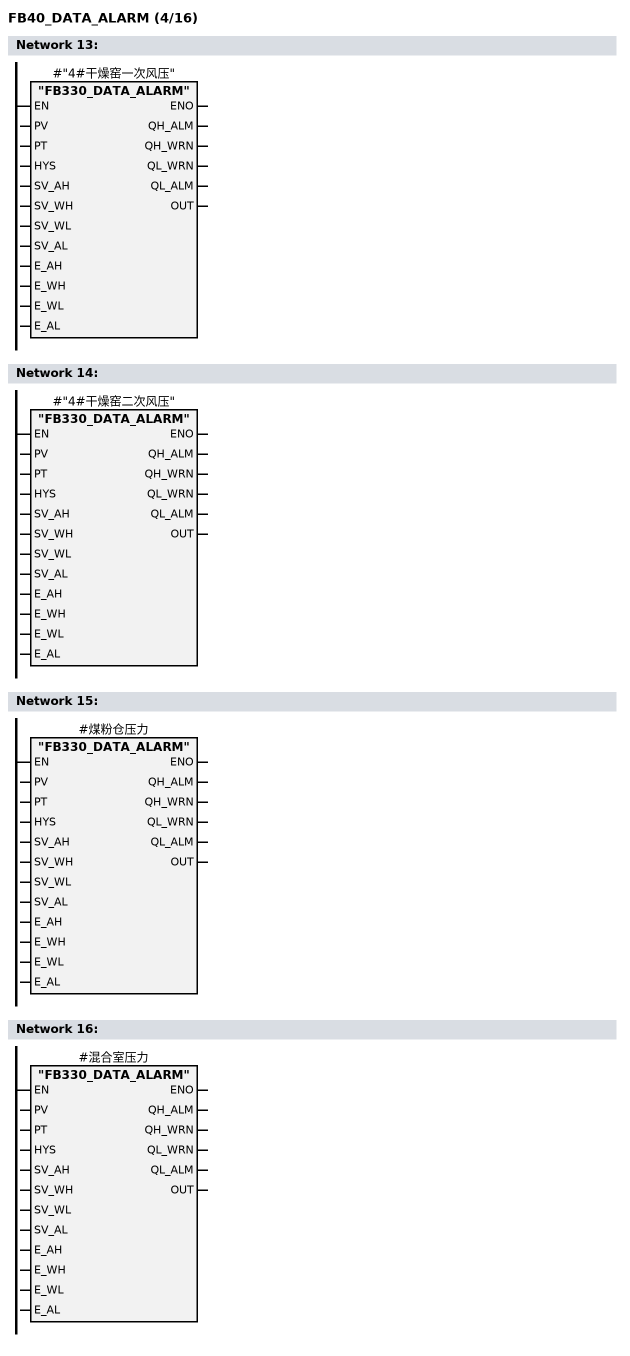
   RUNG wire#powerrail
      #"4#干燥窑一次风压"(PV :=, PT :=, HYS :=, SV_AH :=, SV_WH :=, SV_WL :=, SV_AL :=, E_AH :=, E_WH :=, E_WL :=, E_AL :=, QH_ALM =>, QH_WRN =>, QL_WRN =>, QL_ALM =>, OUT =>)
   END_RUNG
   // the same network as SCL:
   #"4#干燥窑一次风压"();   // "FB330_DATA_ALARM"
END_REGION

REGION Network 14
   RUNG wire#powerrail
      #"4#干燥窑二次风压"(PV :=, PT :=, HYS :=, SV_AH :=, SV_WH :=, SV_WL :=, SV_AL :=, E_AH :=, E_WH :=, E_WL :=, E_AL :=, QH_ALM =>, QH_WRN =>, QL_WRN =>, QL_ALM =>, OUT =>)
   END_RUNG
   // the same network as SCL:
   #"4#干燥窑二次风压"();   // "FB330_DATA_ALARM"
END_REGION

REGION Network 15
   RUNG wire#powerrail
      #煤粉仓压力(PV :=, PT :=, HYS :=, SV_AH :=, SV_WH :=, SV_WL :=, SV_AL :=, E_AH :=, E_WH :=, E_WL :=, E_AL :=, QH_ALM =>, QH_WRN =>, QL_WRN =>, QL_ALM =>, OUT =>)
   END_RUNG
   // the same network as SCL:
   #煤粉仓压力();   // "FB330_DATA_ALARM"
END_REGION

REGION Network 16
   RUNG wire#powerrail
      #混合室压力(PV :=, PT :=, HYS :=, SV_AH :=, SV_WH :=, SV_WL :=, SV_AL :=, E_AH :=, E_WH :=, E_WL :=, E_AL :=, QH_ALM =>, QH_WRN =>, QL_WRN =>, QL_ALM =>, OUT =>)
   END_RUNG
   // the same network as SCL:
   #混合室压力();   // "FB330_DATA_ALARM"
END_REGION

REGION Network 17
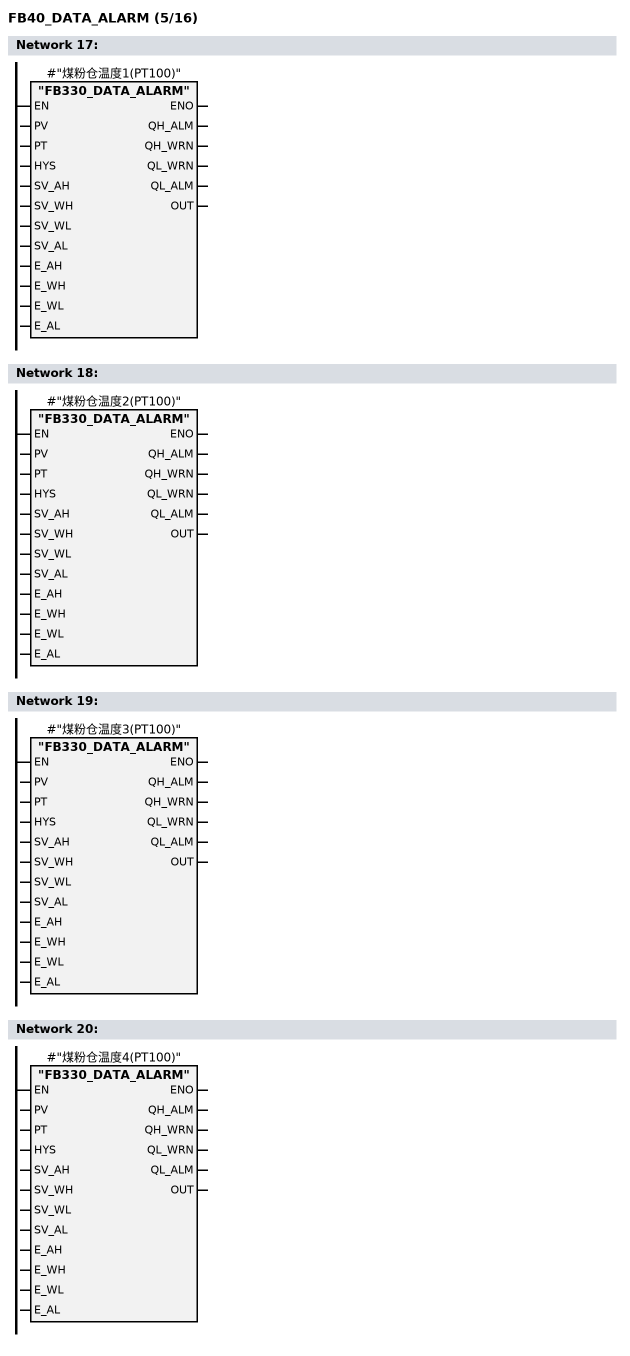
   RUNG wire#powerrail
      #"煤粉仓温度1(PT100)"(PV :=, PT :=, HYS :=, SV_AH :=, SV_WH :=, SV_WL :=, SV_AL :=, E_AH :=, E_WH :=, E_WL :=, E_AL :=, QH_ALM =>, QH_WRN =>, QL_WRN =>, QL_ALM =>, OUT =>)
   END_RUNG
   // the same network as SCL:
   #"煤粉仓温度1(PT100)"();   // "FB330_DATA_ALARM"
END_REGION

REGION Network 18
   RUNG wire#powerrail
      #"煤粉仓温度2(PT100)"(PV :=, PT :=, HYS :=, SV_AH :=, SV_WH :=, SV_WL :=, SV_AL :=, E_AH :=, E_WH :=, E_WL :=, E_AL :=, QH_ALM =>, QH_WRN =>, QL_WRN =>, QL_ALM =>, OUT =>)
   END_RUNG
   // the same network as SCL:
   #"煤粉仓温度2(PT100)"();   // "FB330_DATA_ALARM"
END_REGION

REGION Network 19
   RUNG wire#powerrail
      #"煤粉仓温度3(PT100)"(PV :=, PT :=, HYS :=, SV_AH :=, SV_WH :=, SV_WL :=, SV_AL :=, E_AH :=, E_WH :=, E_WL :=, E_AL :=, QH_ALM =>, QH_WRN =>, QL_WRN =>, QL_ALM =>, OUT =>)
   END_RUNG
   // the same network as SCL:
   #"煤粉仓温度3(PT100)"();   // "FB330_DATA_ALARM"
END_REGION

REGION Network 20
   RUNG wire#powerrail
      #"煤粉仓温度4(PT100)"(PV :=, PT :=, HYS :=, SV_AH :=, SV_WH :=, SV_WL :=, SV_AL :=, E_AH :=, E_WH :=, E_WL :=, E_AL :=, QH_ALM =>, QH_WRN =>, QL_WRN =>, QL_ALM =>, OUT =>)
   END_RUNG
   // the same network as SCL:
   #"煤粉仓温度4(PT100)"();   // "FB330_DATA_ALARM"
END_REGION

REGION Network 21
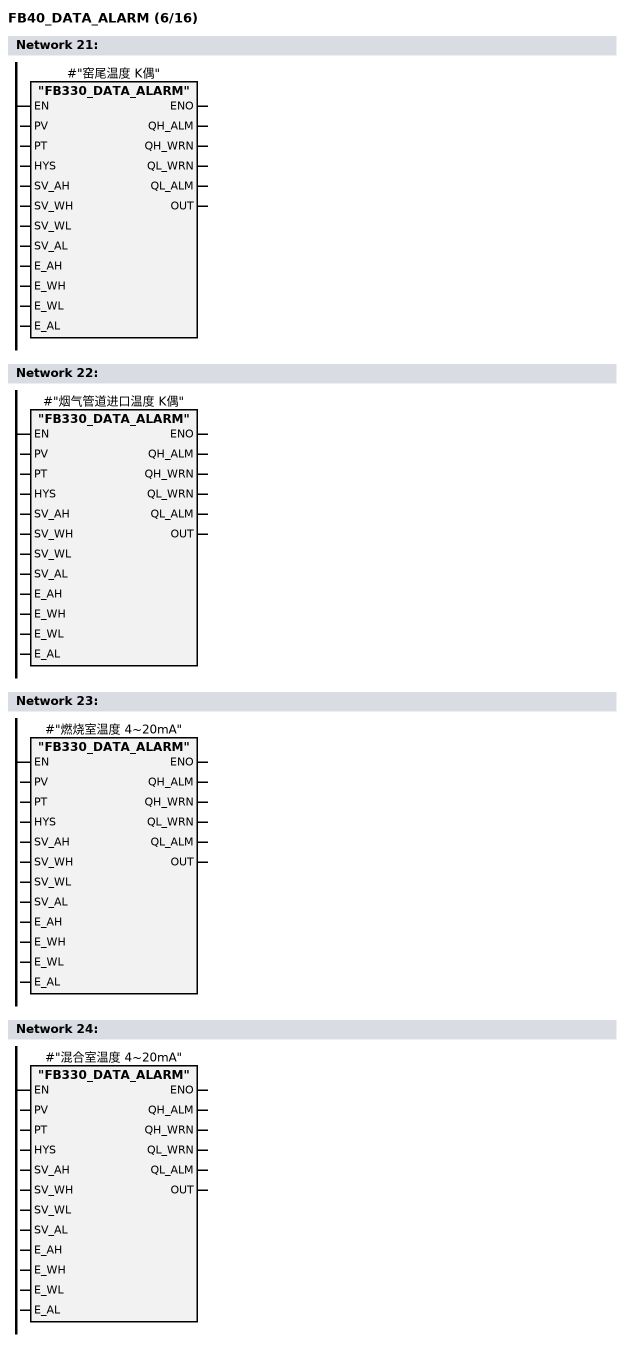
   RUNG wire#powerrail
      #"窑尾温度 K偶"(PV :=, PT :=, HYS :=, SV_AH :=, SV_WH :=, SV_WL :=, SV_AL :=, E_AH :=, E_WH :=, E_WL :=, E_AL :=, QH_ALM =>, QH_WRN =>, QL_WRN =>, QL_ALM =>, OUT =>)
   END_RUNG
   // the same network as SCL:
   #"窑尾温度 K偶"();   // "FB330_DATA_ALARM"
END_REGION

REGION Network 22
   RUNG wire#powerrail
      #"烟气管道进口温度 K偶"(PV :=, PT :=, HYS :=, SV_AH :=, SV_WH :=, SV_WL :=, SV_AL :=, E_AH :=, E_WH :=, E_WL :=, E_AL :=, QH_ALM =>, QH_WRN =>, QL_WRN =>, QL_ALM =>, OUT =>)
   END_RUNG
   // the same network as SCL:
   #"烟气管道进口温度 K偶"();   // "FB330_DATA_ALARM"
END_REGION

REGION Network 23
   RUNG wire#powerrail
      #"燃烧室温度 4~20mA"(PV :=, PT :=, HYS :=, SV_AH :=, SV_WH :=, SV_WL :=, SV_AL :=, E_AH :=, E_WH :=, E_WL :=, E_AL :=, QH_ALM =>, QH_WRN =>, QL_WRN =>, QL_ALM =>, OUT =>)
   END_RUNG
   // the same network as SCL:
   #"燃烧室温度 4~20mA"();   // "FB330_DATA_ALARM"
END_REGION

REGION Network 24
   RUNG wire#powerrail
      #"混合室温度 4~20mA"(PV :=, PT :=, HYS :=, SV_AH :=, SV_WH :=, SV_WL :=, SV_AL :=, E_AH :=, E_WH :=, E_WL :=, E_AL :=, QH_ALM =>, QH_WRN =>, QL_WRN =>, QL_ALM =>, OUT =>)
   END_RUNG
   // the same network as SCL:
   #"混合室温度 4~20mA"();   // "FB330_DATA_ALARM"
END_REGION

REGION Network 25
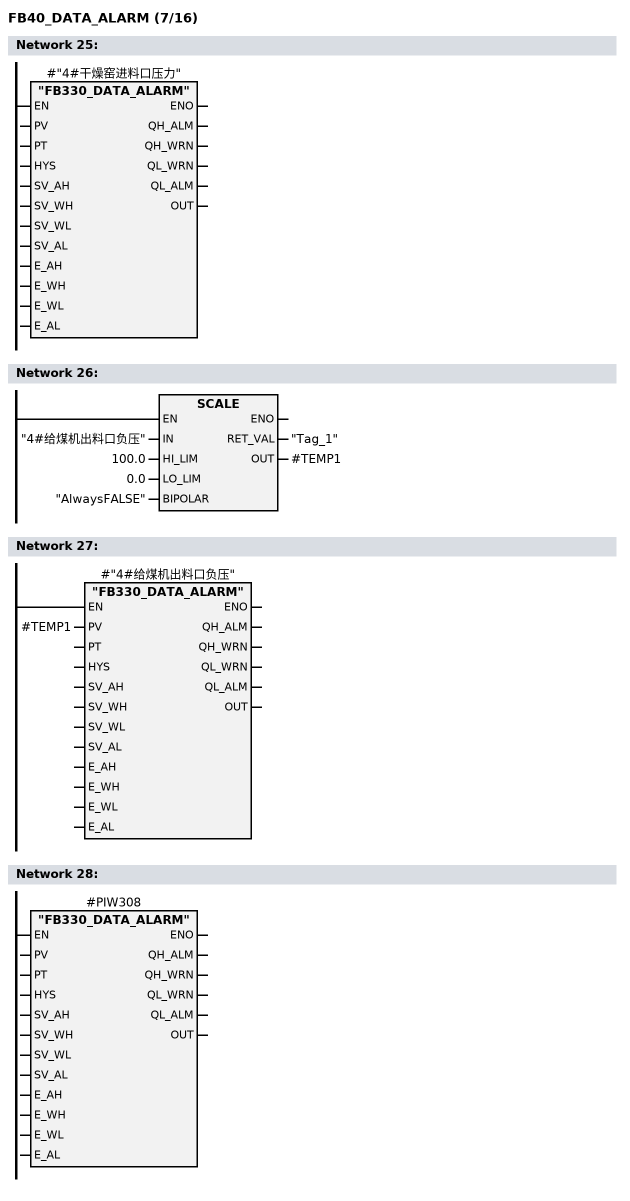
   RUNG wire#powerrail
      #"4#干燥窑进料口压力"(PV :=, PT :=, HYS :=, SV_AH :=, SV_WH :=, SV_WL :=, SV_AL :=, E_AH :=, E_WH :=, E_WL :=, E_AL :=, QH_ALM =>, QH_WRN =>, QL_WRN =>, QL_ALM =>, OUT =>)
   END_RUNG
   // the same network as SCL:
   #"4#干燥窑进料口压力"();   // "FB330_DATA_ALARM"
END_REGION

REGION Network 26
   "Tag_1" := SCALE(IN := "4#给煤机出料口负压", HI_LIM := 100.0, LO_LIM := 0.0, BIPOLAR := "AlwaysFALSE", OUT => #TEMP1);
END_REGION

REGION Network 27
   RUNG wire#powerrail
      #"4#给煤机出料口负压"(PV := #TEMP1, PT :=, HYS :=, SV_AH :=, SV_WH :=, SV_WL :=, SV_AL :=, E_AH :=, E_WH :=, E_WL :=, E_AL :=, QH_ALM =>, QH_WRN =>, QL_WRN =>, QL_ALM =>, OUT =>)
   END_RUNG
   // the same network as SCL:
   #"4#给煤机出料口负压"(PV := #TEMP1);   // "FB330_DATA_ALARM"
END_REGION

REGION Network 28
   RUNG wire#powerrail
      #PIW308(PV :=, PT :=, HYS :=, SV_AH :=, SV_WH :=, SV_WL :=, SV_AL :=, E_AH :=, E_WH :=, E_WL :=, E_AL :=, QH_ALM =>, QH_WRN =>, QL_WRN =>, QL_ALM =>, OUT =>)
   END_RUNG
   // the same network as SCL:
   #PIW308();   // "FB330_DATA_ALARM"
END_REGION

REGION Network 29
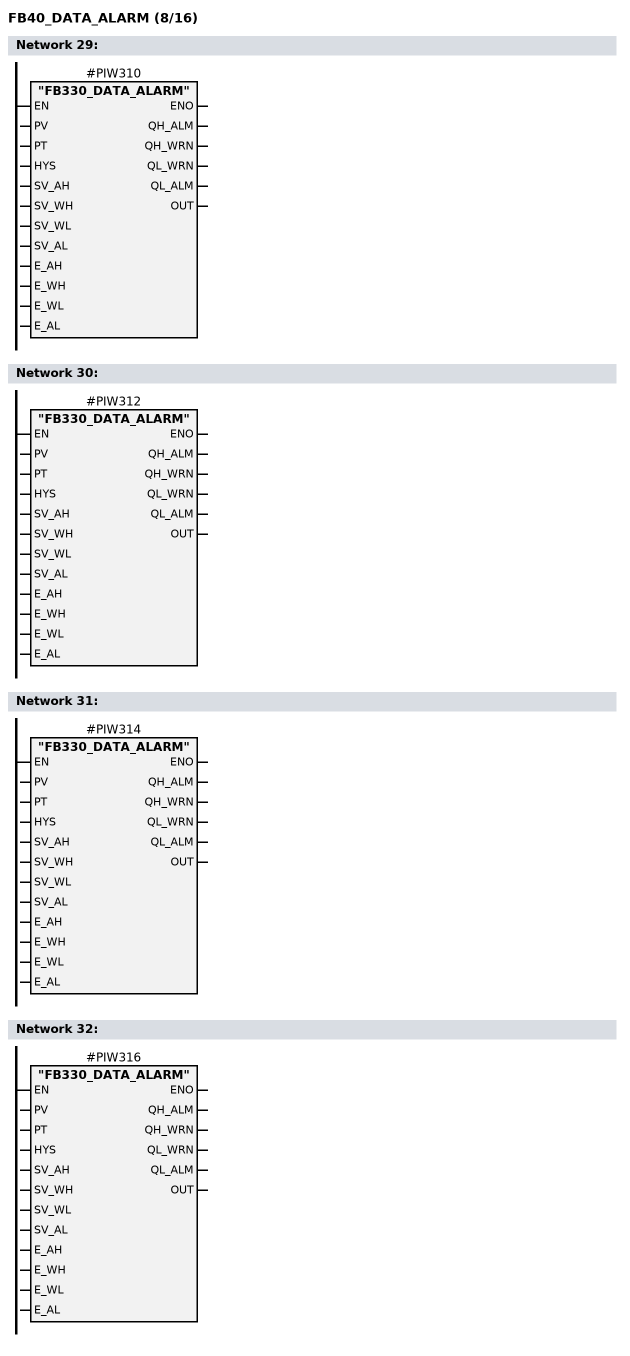
   RUNG wire#powerrail
      #PIW310(PV :=, PT :=, HYS :=, SV_AH :=, SV_WH :=, SV_WL :=, SV_AL :=, E_AH :=, E_WH :=, E_WL :=, E_AL :=, QH_ALM =>, QH_WRN =>, QL_WRN =>, QL_ALM =>, OUT =>)
   END_RUNG
   // the same network as SCL:
   #PIW310();   // "FB330_DATA_ALARM"
END_REGION

REGION Network 30
   RUNG wire#powerrail
      #PIW312(PV :=, PT :=, HYS :=, SV_AH :=, SV_WH :=, SV_WL :=, SV_AL :=, E_AH :=, E_WH :=, E_WL :=, E_AL :=, QH_ALM =>, QH_WRN =>, QL_WRN =>, QL_ALM =>, OUT =>)
   END_RUNG
   // the same network as SCL:
   #PIW312();   // "FB330_DATA_ALARM"
END_REGION

REGION Network 31
   RUNG wire#powerrail
      #PIW314(PV :=, PT :=, HYS :=, SV_AH :=, SV_WH :=, SV_WL :=, SV_AL :=, E_AH :=, E_WH :=, E_WL :=, E_AL :=, QH_ALM =>, QH_WRN =>, QL_WRN =>, QL_ALM =>, OUT =>)
   END_RUNG
   // the same network as SCL:
   #PIW314();   // "FB330_DATA_ALARM"
END_REGION

REGION Network 32
   RUNG wire#powerrail
      #PIW316(PV :=, PT :=, HYS :=, SV_AH :=, SV_WH :=, SV_WL :=, SV_AL :=, E_AH :=, E_WH :=, E_WL :=, E_AL :=, QH_ALM =>, QH_WRN =>, QL_WRN =>, QL_ALM =>, OUT =>)
   END_RUNG
   // the same network as SCL:
   #PIW316();   // "FB330_DATA_ALARM"
END_REGION

REGION Network 33
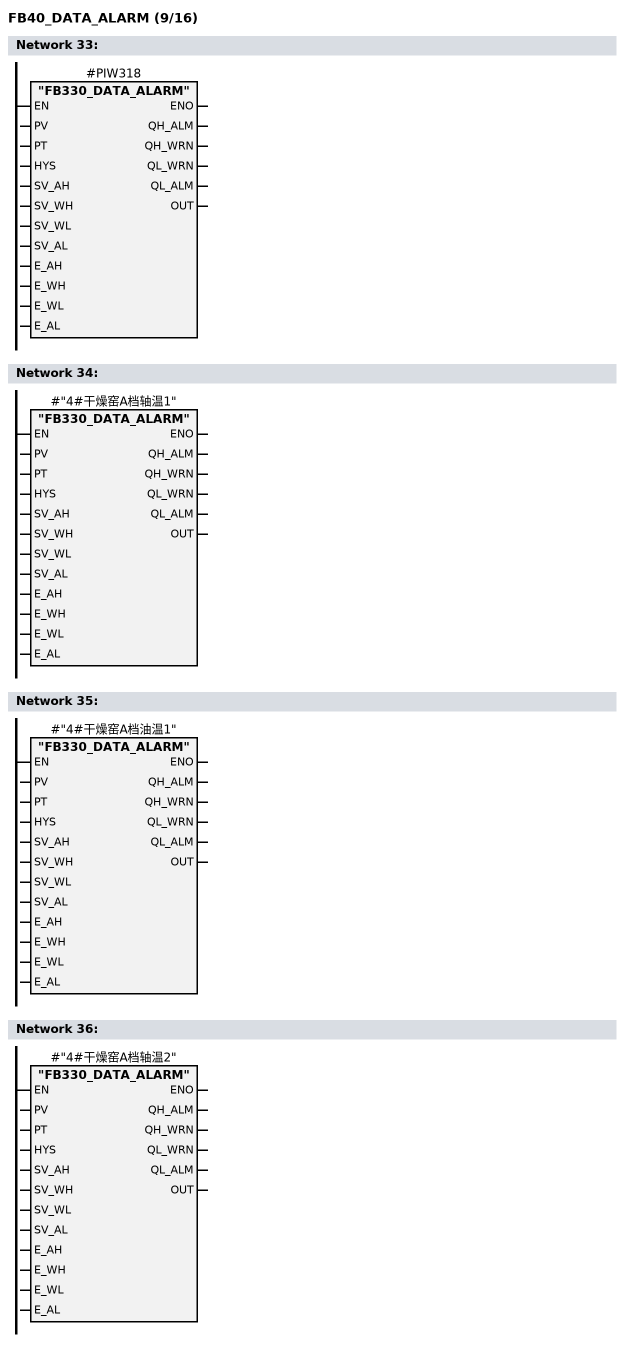
   RUNG wire#powerrail
      #PIW318(PV :=, PT :=, HYS :=, SV_AH :=, SV_WH :=, SV_WL :=, SV_AL :=, E_AH :=, E_WH :=, E_WL :=, E_AL :=, QH_ALM =>, QH_WRN =>, QL_WRN =>, QL_ALM =>, OUT =>)
   END_RUNG
   // the same network as SCL:
   #PIW318();   // "FB330_DATA_ALARM"
END_REGION

REGION Network 34
   RUNG wire#powerrail
      #"4#干燥窑A档轴温1"(PV :=, PT :=, HYS :=, SV_AH :=, SV_WH :=, SV_WL :=, SV_AL :=, E_AH :=, E_WH :=, E_WL :=, E_AL :=, QH_ALM =>, QH_WRN =>, QL_WRN =>, QL_ALM =>, OUT =>)
   END_RUNG
   // the same network as SCL:
   #"4#干燥窑A档轴温1"();   // "FB330_DATA_ALARM"
END_REGION

REGION Network 35
   RUNG wire#powerrail
      #"4#干燥窑A档油温1"(PV :=, PT :=, HYS :=, SV_AH :=, SV_WH :=, SV_WL :=, SV_AL :=, E_AH :=, E_WH :=, E_WL :=, E_AL :=, QH_ALM =>, QH_WRN =>, QL_WRN =>, QL_ALM =>, OUT =>)
   END_RUNG
   // the same network as SCL:
   #"4#干燥窑A档油温1"();   // "FB330_DATA_ALARM"
END_REGION

REGION Network 36
   RUNG wire#powerrail
      #"4#干燥窑A档轴温2"(PV :=, PT :=, HYS :=, SV_AH :=, SV_WH :=, SV_WL :=, SV_AL :=, E_AH :=, E_WH :=, E_WL :=, E_AL :=, QH_ALM =>, QH_WRN =>, QL_WRN =>, QL_ALM =>, OUT =>)
   END_RUNG
   // the same network as SCL:
   #"4#干燥窑A档轴温2"();   // "FB330_DATA_ALARM"
END_REGION

REGION Network 37
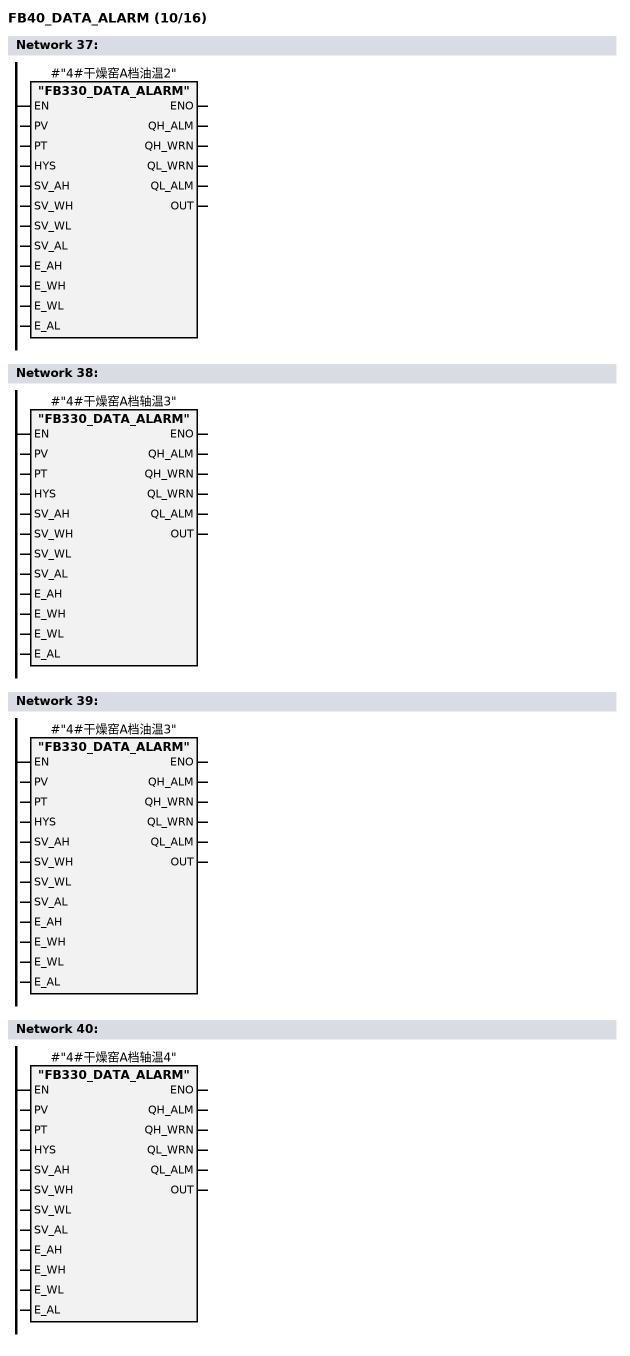
   RUNG wire#powerrail
      #"4#干燥窑A档油温2"(PV :=, PT :=, HYS :=, SV_AH :=, SV_WH :=, SV_WL :=, SV_AL :=, E_AH :=, E_WH :=, E_WL :=, E_AL :=, QH_ALM =>, QH_WRN =>, QL_WRN =>, QL_ALM =>, OUT =>)
   END_RUNG
   // the same network as SCL:
   #"4#干燥窑A档油温2"();   // "FB330_DATA_ALARM"
END_REGION

REGION Network 38
   RUNG wire#powerrail
      #"4#干燥窑A档轴温3"(PV :=, PT :=, HYS :=, SV_AH :=, SV_WH :=, SV_WL :=, SV_AL :=, E_AH :=, E_WH :=, E_WL :=, E_AL :=, QH_ALM =>, QH_WRN =>, QL_WRN =>, QL_ALM =>, OUT =>)
   END_RUNG
   // the same network as SCL:
   #"4#干燥窑A档轴温3"();   // "FB330_DATA_ALARM"
END_REGION

REGION Network 39
   RUNG wire#powerrail
      #"4#干燥窑A档油温3"(PV :=, PT :=, HYS :=, SV_AH :=, SV_WH :=, SV_WL :=, SV_AL :=, E_AH :=, E_WH :=, E_WL :=, E_AL :=, QH_ALM =>, QH_WRN =>, QL_WRN =>, QL_ALM =>, OUT =>)
   END_RUNG
   // the same network as SCL:
   #"4#干燥窑A档油温3"();   // "FB330_DATA_ALARM"
END_REGION

REGION Network 40
   RUNG wire#powerrail
      #"4#干燥窑A档轴温4"(PV :=, PT :=, HYS :=, SV_AH :=, SV_WH :=, SV_WL :=, SV_AL :=, E_AH :=, E_WH :=, E_WL :=, E_AL :=, QH_ALM =>, QH_WRN =>, QL_WRN =>, QL_ALM =>, OUT =>)
   END_RUNG
   // the same network as SCL:
   #"4#干燥窑A档轴温4"();   // "FB330_DATA_ALARM"
END_REGION

REGION Network 41
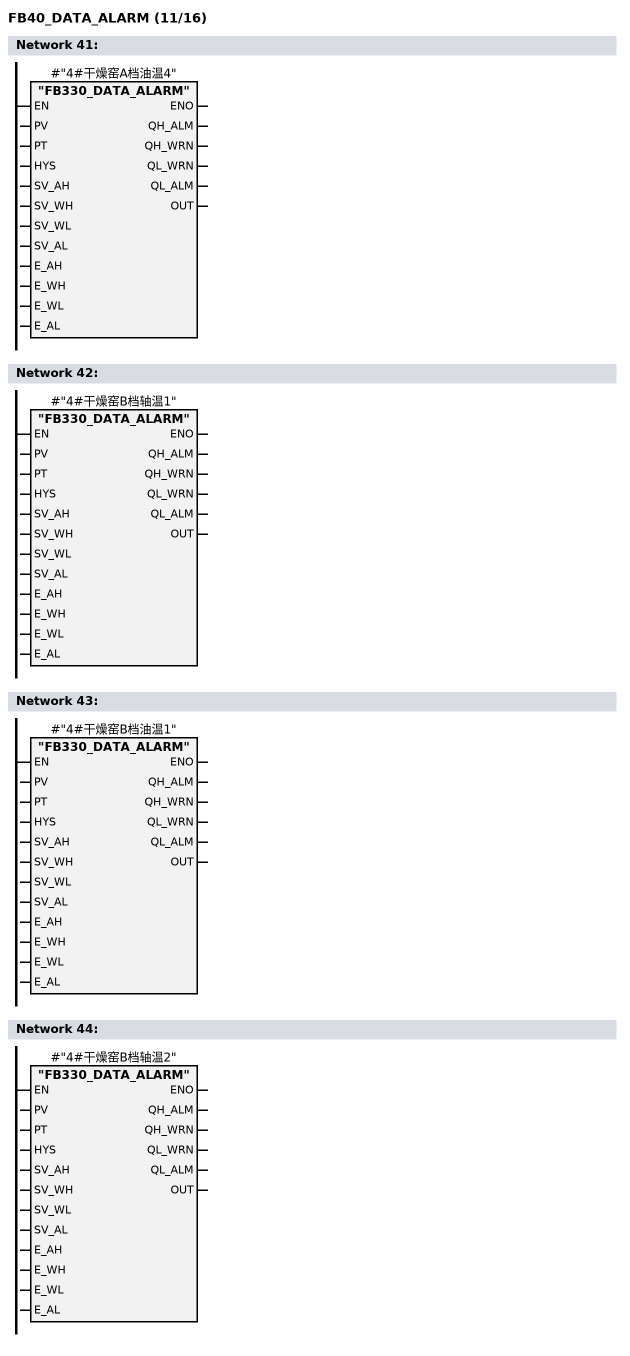
   RUNG wire#powerrail
      #"4#干燥窑A档油温4"(PV :=, PT :=, HYS :=, SV_AH :=, SV_WH :=, SV_WL :=, SV_AL :=, E_AH :=, E_WH :=, E_WL :=, E_AL :=, QH_ALM =>, QH_WRN =>, QL_WRN =>, QL_ALM =>, OUT =>)
   END_RUNG
   // the same network as SCL:
   #"4#干燥窑A档油温4"();   // "FB330_DATA_ALARM"
END_REGION

REGION Network 42
   RUNG wire#powerrail
      #"4#干燥窑B档轴温1"(PV :=, PT :=, HYS :=, SV_AH :=, SV_WH :=, SV_WL :=, SV_AL :=, E_AH :=, E_WH :=, E_WL :=, E_AL :=, QH_ALM =>, QH_WRN =>, QL_WRN =>, QL_ALM =>, OUT =>)
   END_RUNG
   // the same network as SCL:
   #"4#干燥窑B档轴温1"();   // "FB330_DATA_ALARM"
END_REGION

REGION Network 43
   RUNG wire#powerrail
      #"4#干燥窑B档油温1"(PV :=, PT :=, HYS :=, SV_AH :=, SV_WH :=, SV_WL :=, SV_AL :=, E_AH :=, E_WH :=, E_WL :=, E_AL :=, QH_ALM =>, QH_WRN =>, QL_WRN =>, QL_ALM =>, OUT =>)
   END_RUNG
   // the same network as SCL:
   #"4#干燥窑B档油温1"();   // "FB330_DATA_ALARM"
END_REGION

REGION Network 44
   RUNG wire#powerrail
      #"4#干燥窑B档轴温2"(PV :=, PT :=, HYS :=, SV_AH :=, SV_WH :=, SV_WL :=, SV_AL :=, E_AH :=, E_WH :=, E_WL :=, E_AL :=, QH_ALM =>, QH_WRN =>, QL_WRN =>, QL_ALM =>, OUT =>)
   END_RUNG
   // the same network as SCL:
   #"4#干燥窑B档轴温2"();   // "FB330_DATA_ALARM"
END_REGION

REGION Network 45
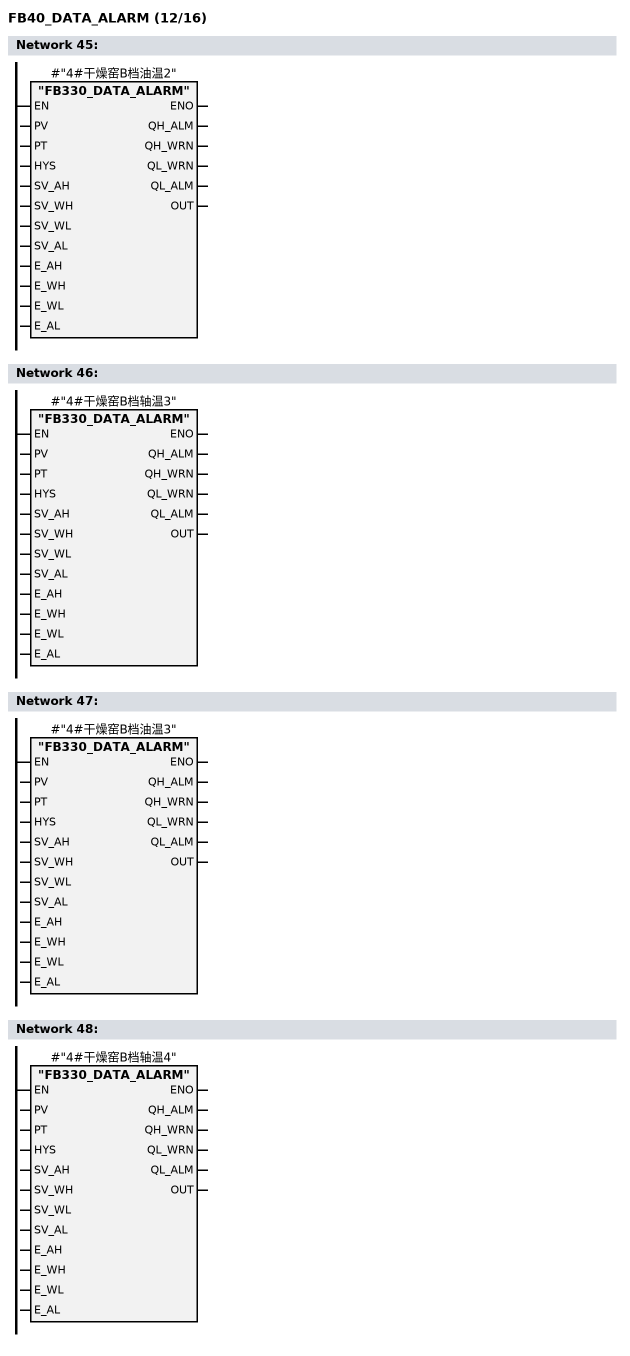
   RUNG wire#powerrail
      #"4#干燥窑B档油温2"(PV :=, PT :=, HYS :=, SV_AH :=, SV_WH :=, SV_WL :=, SV_AL :=, E_AH :=, E_WH :=, E_WL :=, E_AL :=, QH_ALM =>, QH_WRN =>, QL_WRN =>, QL_ALM =>, OUT =>)
   END_RUNG
   // the same network as SCL:
   #"4#干燥窑B档油温2"();   // "FB330_DATA_ALARM"
END_REGION

REGION Network 46
   RUNG wire#powerrail
      #"4#干燥窑B档轴温3"(PV :=, PT :=, HYS :=, SV_AH :=, SV_WH :=, SV_WL :=, SV_AL :=, E_AH :=, E_WH :=, E_WL :=, E_AL :=, QH_ALM =>, QH_WRN =>, QL_WRN =>, QL_ALM =>, OUT =>)
   END_RUNG
   // the same network as SCL:
   #"4#干燥窑B档轴温3"();   // "FB330_DATA_ALARM"
END_REGION

REGION Network 47
   RUNG wire#powerrail
      #"4#干燥窑B档油温3"(PV :=, PT :=, HYS :=, SV_AH :=, SV_WH :=, SV_WL :=, SV_AL :=, E_AH :=, E_WH :=, E_WL :=, E_AL :=, QH_ALM =>, QH_WRN =>, QL_WRN =>, QL_ALM =>, OUT =>)
   END_RUNG
   // the same network as SCL:
   #"4#干燥窑B档油温3"();   // "FB330_DATA_ALARM"
END_REGION

REGION Network 48
   RUNG wire#powerrail
      #"4#干燥窑B档轴温4"(PV :=, PT :=, HYS :=, SV_AH :=, SV_WH :=, SV_WL :=, SV_AL :=, E_AH :=, E_WH :=, E_WL :=, E_AL :=, QH_ALM =>, QH_WRN =>, QL_WRN =>, QL_ALM =>, OUT =>)
   END_RUNG
   // the same network as SCL:
   #"4#干燥窑B档轴温4"();   // "FB330_DATA_ALARM"
END_REGION

REGION Network 49
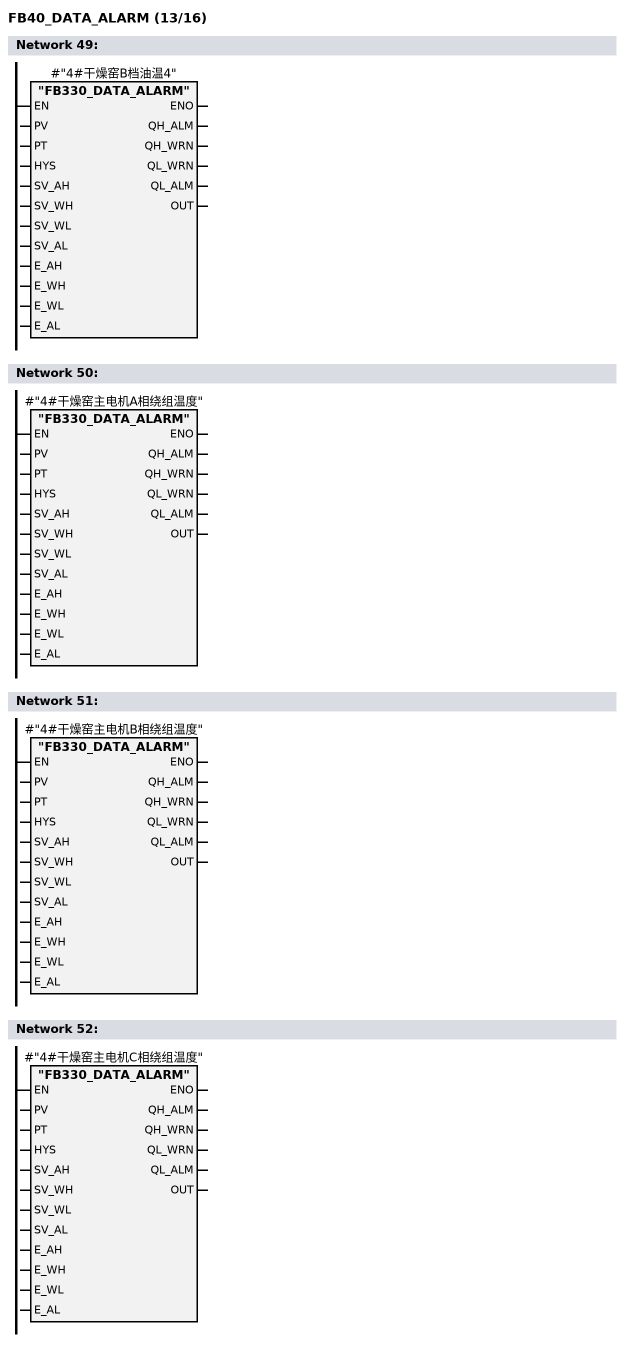
   RUNG wire#powerrail
      #"4#干燥窑B档油温4"(PV :=, PT :=, HYS :=, SV_AH :=, SV_WH :=, SV_WL :=, SV_AL :=, E_AH :=, E_WH :=, E_WL :=, E_AL :=, QH_ALM =>, QH_WRN =>, QL_WRN =>, QL_ALM =>, OUT =>)
   END_RUNG
   // the same network as SCL:
   #"4#干燥窑B档油温4"();   // "FB330_DATA_ALARM"
END_REGION

REGION Network 50
   RUNG wire#powerrail
      #"4#干燥窑主电机A相绕组温度"(PV :=, PT :=, HYS :=, SV_AH :=, SV_WH :=, SV_WL :=, SV_AL :=, E_AH :=, E_WH :=, E_WL :=, E_AL :=, QH_ALM =>, QH_WRN =>, QL_WRN =>, QL_ALM =>, OUT =>)
   END_RUNG
   // the same network as SCL:
   #"4#干燥窑主电机A相绕组温度"();   // "FB330_DATA_ALARM"
END_REGION

REGION Network 51
   RUNG wire#powerrail
      #"4#干燥窑主电机B相绕组温度"(PV :=, PT :=, HYS :=, SV_AH :=, SV_WH :=, SV_WL :=, SV_AL :=, E_AH :=, E_WH :=, E_WL :=, E_AL :=, QH_ALM =>, QH_WRN =>, QL_WRN =>, QL_ALM =>, OUT =>)
   END_RUNG
   // the same network as SCL:
   #"4#干燥窑主电机B相绕组温度"();   // "FB330_DATA_ALARM"
END_REGION

REGION Network 52
   RUNG wire#powerrail
      #"4#干燥窑主电机C相绕组温度"(PV :=, PT :=, HYS :=, SV_AH :=, SV_WH :=, SV_WL :=, SV_AL :=, E_AH :=, E_WH :=, E_WL :=, E_AL :=, QH_ALM =>, QH_WRN =>, QL_WRN =>, QL_ALM =>, OUT =>)
   END_RUNG
   // the same network as SCL:
   #"4#干燥窑主电机C相绕组温度"();   // "FB330_DATA_ALARM"
END_REGION

REGION Network 53
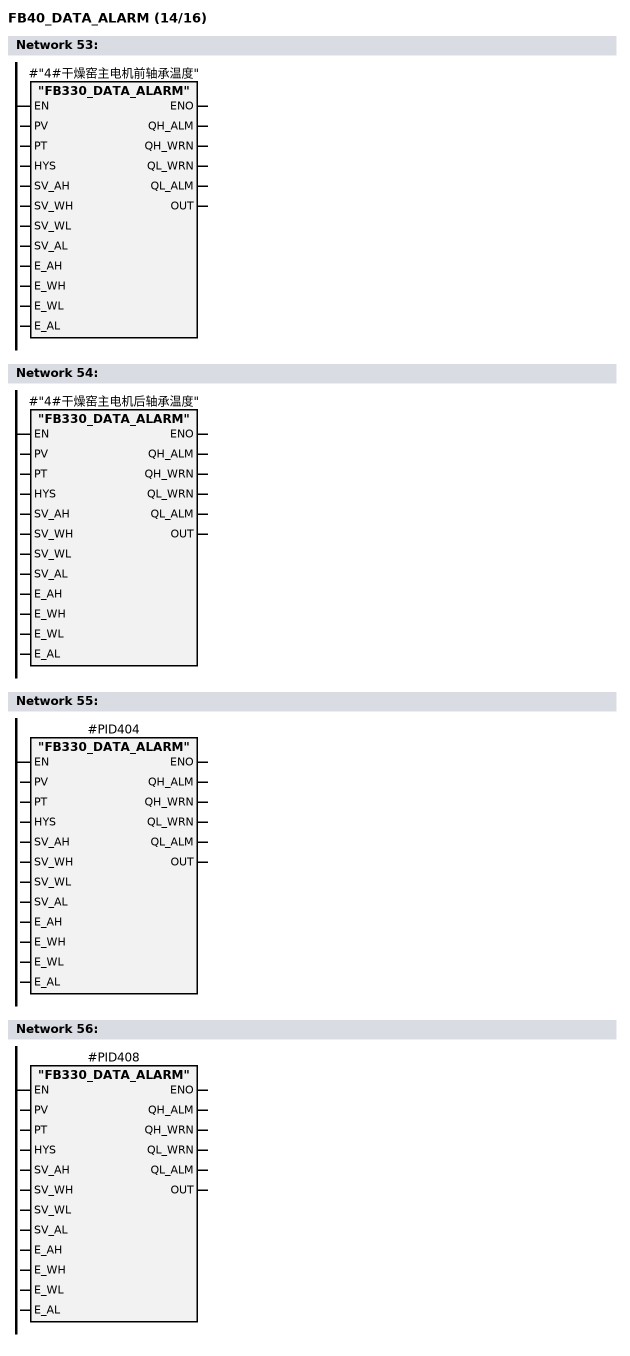
   RUNG wire#powerrail
      #"4#干燥窑主电机前轴承温度"(PV :=, PT :=, HYS :=, SV_AH :=, SV_WH :=, SV_WL :=, SV_AL :=, E_AH :=, E_WH :=, E_WL :=, E_AL :=, QH_ALM =>, QH_WRN =>, QL_WRN =>, QL_ALM =>, OUT =>)
   END_RUNG
   // the same network as SCL:
   #"4#干燥窑主电机前轴承温度"();   // "FB330_DATA_ALARM"
END_REGION

REGION Network 54
   RUNG wire#powerrail
      #"4#干燥窑主电机后轴承温度"(PV :=, PT :=, HYS :=, SV_AH :=, SV_WH :=, SV_WL :=, SV_AL :=, E_AH :=, E_WH :=, E_WL :=, E_AL :=, QH_ALM =>, QH_WRN =>, QL_WRN =>, QL_ALM =>, OUT =>)
   END_RUNG
   // the same network as SCL:
   #"4#干燥窑主电机后轴承温度"();   // "FB330_DATA_ALARM"
END_REGION

REGION Network 55
   RUNG wire#powerrail
      #PID404(PV :=, PT :=, HYS :=, SV_AH :=, SV_WH :=, SV_WL :=, SV_AL :=, E_AH :=, E_WH :=, E_WL :=, E_AL :=, QH_ALM =>, QH_WRN =>, QL_WRN =>, QL_ALM =>, OUT =>)
   END_RUNG
   // the same network as SCL:
   #PID404();   // "FB330_DATA_ALARM"
END_REGION

REGION Network 56
   RUNG wire#powerrail
      #PID408(PV :=, PT :=, HYS :=, SV_AH :=, SV_WH :=, SV_WL :=, SV_AL :=, E_AH :=, E_WH :=, E_WL :=, E_AL :=, QH_ALM =>, QH_WRN =>, QL_WRN =>, QL_ALM =>, OUT =>)
   END_RUNG
   // the same network as SCL:
   #PID408();   // "FB330_DATA_ALARM"
END_REGION

REGION Network 57
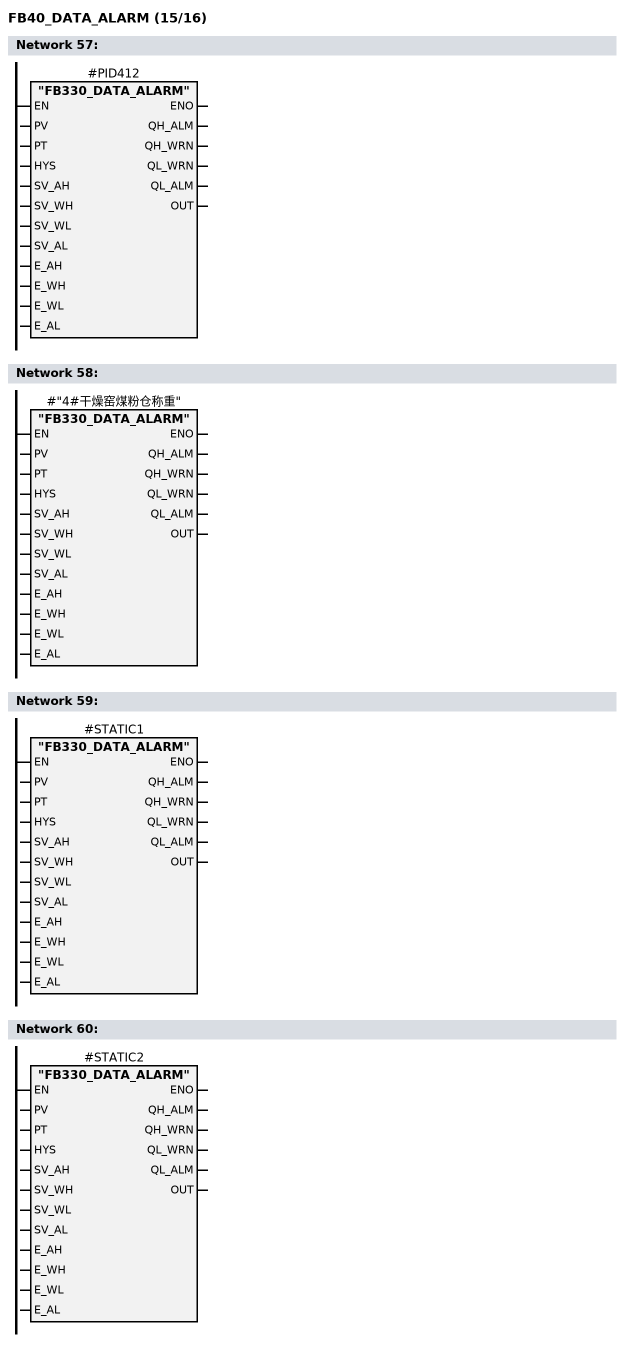
   RUNG wire#powerrail
      #PID412(PV :=, PT :=, HYS :=, SV_AH :=, SV_WH :=, SV_WL :=, SV_AL :=, E_AH :=, E_WH :=, E_WL :=, E_AL :=, QH_ALM =>, QH_WRN =>, QL_WRN =>, QL_ALM =>, OUT =>)
   END_RUNG
   // the same network as SCL:
   #PID412();   // "FB330_DATA_ALARM"
END_REGION

REGION Network 58
   RUNG wire#powerrail
      #"4#干燥窑煤粉仓称重"(PV :=, PT :=, HYS :=, SV_AH :=, SV_WH :=, SV_WL :=, SV_AL :=, E_AH :=, E_WH :=, E_WL :=, E_AL :=, QH_ALM =>, QH_WRN =>, QL_WRN =>, QL_ALM =>, OUT =>)
   END_RUNG
   // the same network as SCL:
   #"4#干燥窑煤粉仓称重"();   // "FB330_DATA_ALARM"
END_REGION

REGION Network 59
   RUNG wire#powerrail
      #STATIC1(PV :=, PT :=, HYS :=, SV_AH :=, SV_WH :=, SV_WL :=, SV_AL :=, E_AH :=, E_WH :=, E_WL :=, E_AL :=, QH_ALM =>, QH_WRN =>, QL_WRN =>, QL_ALM =>, OUT =>)
   END_RUNG
   // the same network as SCL:
   #STATIC1();   // "FB330_DATA_ALARM"
END_REGION

REGION Network 60
   RUNG wire#powerrail
      #STATIC2(PV :=, PT :=, HYS :=, SV_AH :=, SV_WH :=, SV_WL :=, SV_AL :=, E_AH :=, E_WH :=, E_WL :=, E_AL :=, QH_ALM =>, QH_WRN =>, QL_WRN =>, QL_ALM =>, OUT =>)
   END_RUNG
   // the same network as SCL:
   #STATIC2();   // "FB330_DATA_ALARM"
END_REGION

REGION Network 61
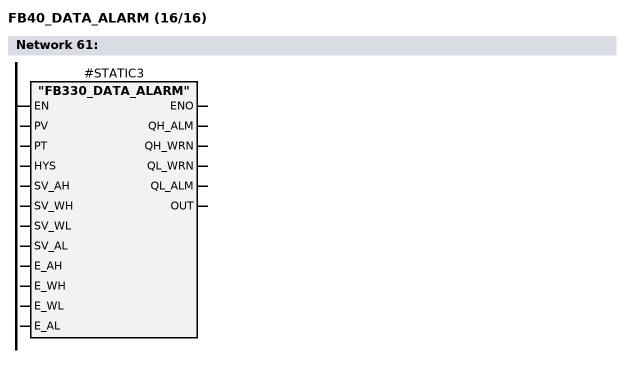
   RUNG wire#powerrail
      #STATIC3(PV :=, PT :=, HYS :=, SV_AH :=, SV_WH :=, SV_WL :=, SV_AL :=, E_AH :=, E_WH :=, E_WL :=, E_AL :=, QH_ALM =>, QH_WRN =>, QL_WRN =>, QL_ALM =>, OUT =>)
   END_RUNG
   // the same network as SCL:
   #STATIC3();   // "FB330_DATA_ALARM"
END_REGION
END_FUNCTION_BLOCK

FUNCTION_BLOCK "FB330_DATA_ALARM"   // FB330, LAD
{ S7_Optimized_Access := 'FALSE' }
VERSION : 0.1
// REAL的报警块
   VAR_INPUT
      PV : Real;   // 过程值
      PT : Real := 1.0;   // 系数
      HYS : Real;   // 回差值
      SV_AH : Real;   // 高报警设定值
      SV_WH : Real;   // 高警告设定值
      SV_WL : Real;   // 低警告设定值
      SV_AL : Real;   // 低报警设定值
      E_AH : Bool;   // 高报警使能
      E_WH : Bool;   // 高警告使能
      E_WL : Bool;   // 低警告使能
      E_AL : Bool;   // 低报警使能
   END_VAR
   VAR_OUTPUT
      QH_ALM : Bool;   // 高报警输出
      QH_WRN : Bool;   // 高警告输出
      QL_WRN : Bool;   // 低警告输出
      QL_ALM : Bool;   // 低报警输出
      OUT : Real;   // 输出
   END_VAR
   VAR
      SR1 : Bool;
      SR2 : Bool;
      SR3 : Bool;
      SR4 : Bool;
   END_VAR
   VAR_TEMP
      TEMP_AH : Real;
      TEMP_WH : Real;
      TEMP_AL : Real;
      TEMP_WL : Real;
      TEMP_OUT : Real;
   END_VAR
BEGIN
